   "DB611_Hydraulic_State_MH_Hydraulic{2}_Switch_Hydraulic_ON_OFF" : Bool = PLC DB939_Tool_alloc_HMI.SaveSortProg_name[7] AT %DB611.DBX26.3, 1 s
   "DB619_State_MPart_Recirculation{2}_Switch_Intervall" : Bool = PLC DB619_State_MPart.Recirculation[2].Switch_Intervall AT %DB619.DBX72.0, 1 s
   "DB619_State_MPart_Recirculation{2}_Switch_Lowpressure" : Bool = PLC DB619_State_MPart.Recirculation[2].Switch_Lowpressure AT %DB619.DBX72.2, 1 s
   "DB619_State_MPart_Recirculation{2}_Switch_Reduced" : Bool = PLC DB619_State_MPart.Recirculation[2].Switch_Reduced AT %DB619.DBX72.3, 1 s
   "DB619_State_MPart_Recirculation{2}_State_Intervall" : Int = PLC DB619_State_MPart.Recirculation[2].State_Intervall AT %DB619.DBW74, 1 s
   "DB619_State_MPart_Recirculation{2}_State_Lowpressure" : Int = PLC DB619_State_MPart.Recirculation[2].State_Lowpressure AT %DB619.DBW76, 1 s
   "DB619_State_MPart_Recirculation{2}_State_Reduced" : Int = PLC DB619_State_MPart.Recirculation[2].State_Reduced AT %DB619.DBW78, 1 s

HMI tags "General Machine Configuration"
   "DB790_PlantParameter_AmountMH" : Int = PLC DB790_PlantParameter.AmountMH AT %DB790.DBW4, 1 s
   "DB790_PlantParameter_AmountTank" : Int = PLC DB790_PlantParameter.AmountTank AT %DB790.DBW6, 1 s
   "DB790_PlantParameter_AmountToolStation" : Int = PLC DB790_PlantParameter.AmountToolStation AT %DB790.DBW10, 1 s
   "DB790_PlantParameter_AmountMouldCarrier" : Int = PLC DB790_PlantParameter.AmountMouldCarrier AT %DB790.DBW12, 1 s
   "DB790_PlantParameter_AmountProCanModul" : Int = PLC DB790_PlantParameter.AmountProCanModul AT %DB790.DBW2, 1 s
   "DB790_PlantParameter_AmountMeteringUnits" : Int = PLC DB790_PlantParameter.AmountMeteringUnits AT %DB790.DBW8, 1 s
   "DB790_PlantParameter_AmountMachine" : Int = PLC DB790_PlantParameter.AmountMachine AT %DB790.DBW24, 1 s
   "DB790_PlantParameter_Bit_ProgrammNofromInterface" : Bool = PLC DB790_PlantParameter.Bit.ProgrammNofromInterface AT %DB790.DBX0.3, 1 s
   "DB790_PlantParameter_Bit_MHNofromInterface" : Bool = PLC DB790_PlantParameter.Bit.MHNofromInterface AT %DB790.DBX0.2, 1 s
   "DB790_PlantParameter_AmountRobots" : Int = PLC DB790_PlantParameter.AmountRobots AT %DB790.DBW26, 1 s

HMI tags "Pump"
   "DB608_PV_Metering_Metering{0}_MixingRatio_PV_SetV_WarningLowerLimit" : Real = PLC DB608_PV_Metering.Metering[0].MixingRatio.PV_SetV.WarningLowerLimit AT %DB608.DBD202, 1 s
      on ChangeValue: SetBit("DB608_PV_Metering_Write")
   "DB608_PV_Metering_Metering{0}_MixingRatio_PV_SetV_WarningUpperLimit" : Real = PLC DB608_PV_Metering.Metering[0].MixingRatio.PV_SetV.WarningUpperLimit AT %DB608.DBD206, 1 s
      on ChangeValue: SetBit("DB608_PV_Metering_Write")
   "DB608_PV_Metering_Metering{0}_MixingRatio_PV_SetV_AlarmLowerLimit" : Real = PLC DB608_PV_Metering.Metering[0].MixingRatio.PV_SetV.AlarmLowerLimit AT %DB608.DBD210, 1 s
      on ChangeValue: SetBit("DB608_PV_Metering_Write")
   "DB608_PV_Metering_Metering{0}_MixingRatio_PV_SetV_AlarmUpperLimit" : Real = PLC DB608_PV_Metering.Metering[0].MixingRatio.PV_SetV.AlarmUpperLimit AT %DB608.DBD214, 1 s
      on ChangeValue: SetBit("DB608_PV_Metering_Write")
   "DB608_PV_Metering_Metering{0}_MixingRatio_PV_SetV_Value" : Real = PLC DB608_PV_Metering.Metering[0].MixingRatio.PV_SetV.Value AT %DB608.DBD198, 1 s
      on ChangeValue: SetBit("DB608_PV_Metering_Write")
   "DB608_PV_Metering_Metering{0}_Flow_PV_SetV_Value" : Real = PLC DB608_PV_Metering.Metering[0].Flow.PV_SetV.Value AT %DB608.DBD6, 1 s
      on ChangeValue: SetBit("DB608_PV_Metering_Write")
   "DB608_PV_Metering_Metering{0}_Flow_PV_SetV_WarningLowerLimit" : Real = PLC DB608_PV_Metering.Metering[0].Flow.PV_SetV.WarningLowerLimit AT %DB608.DBD10, 1 s
      on ChangeValue: SetBit("DB608_PV_Metering_Write")
   "DB608_PV_Metering_Metering{0}_Flow_PV_SetV_WarningUpperLimit" : Real = PLC DB608_PV_Metering.Metering[0].Flow.PV_SetV.WarningUpperLimit AT %DB608.DBD14, 1 s
      on ChangeValue: SetBit("DB608_PV_Metering_Write")
   "DB608_PV_Metering_Metering{0}_Flow_PV_SetV_AlarmLowerLimit" : Real = PLC DB608_PV_Metering.Metering[0].Flow.PV_SetV.AlarmLowerLimit AT %DB608.DBD18, 1 s
      on ChangeValue: SetBit("DB608_PV_Metering_Write")
   "DB608_PV_Metering_Metering{0}_Flow_PV_SetV_AlarmUpperLimit" : Real = PLC DB608_PV_Metering.Metering[0].Flow.PV_SetV.AlarmUpperLimit AT %DB608.DBD22, 1 s
      on ChangeValue: SetBit("DB608_PV_Metering_Write")
   "DB608_PV_Metering_Metering{0}_Pressure_PV_SetV_Value" : Real = PLC DB608_PV_Metering.Metering[0].Pressure.PV_SetV.Value AT %DB608.DBD54, 1 s
      on ChangeValue: SetBit("DB608_PV_Metering_Write")
   "DB608_PV_Metering_Metering{0}_Pressure_PV_SetV_WarningLowerLimit" : Real = PLC DB608_PV_Metering.Metering[0].Pressure.PV_SetV.WarningLowerLimit AT %DB608.DBD58, 1 s
      on ChangeValue: SetBit("DB608_PV_Metering_Write")
   "DB608_PV_Metering_Metering{0}_Pressure_PV_SetV_WarningUpperLimit" : Real = PLC DB608_PV_Metering.Metering[0].Pressure.PV_SetV.WarningUpperLimit AT %DB608.DBD62, 1 s
      on ChangeValue: SetBit("DB608_PV_Metering_Write")
   "DB608_PV_Metering_Metering{0}_Pressure_PV_SetV_AlarmLowerLimit" : Real = PLC DB608_PV_Metering.Metering[0].Pressure.PV_SetV.AlarmLowerLimit AT %DB608.DBD66, 1 s
      on ChangeValue: SetBit("DB608_PV_Metering_Write")
   "DB608_PV_Metering_Metering{0}_Pressure_PV_SetV_AlarmUpperLimit" : Real = PLC DB608_PV_Metering.Metering[0].Pressure.PV_SetV.AlarmUpperLimit AT %DB608.DBD70, 1 s
      on ChangeValue: SetBit("DB608_PV_Metering_Write")
   "Metering Display Open" : Int AT %DB1.DBD0
   "DB613_Komponent_State_Read" : Bool = PLC DB613_Komponent_State.Read AT %DB613.DBX6.0, 1 s
   "DB608_PV_Metering_Write" : Bool = PLC DB608_PV_Metering.Write AT %DB608.DBX4.1, 1 s
   "DB613_Komponent_State_ReadDeviceNo" : Int = PLC DB613_Komponent_State.ReadDeviceNo AT %DB613.DBW0, 1 s
      on ChangeValue: SetBit("DB613_Komponent_State_Write")
   "Control" : Int AT %DB1.DBW0
   "DB753_MeteringPump_Pump{0}_MachineNumber" : Byte = PLC DB753_MeteringPump.Pump[0].MachineNumber AT %DB753.DBB25, 1 s
      on ChangeValue: SetBit("DB613_Komponent_State_Write")
   "DB753_MeteringPump_Pump{0}_Name" : String[20] = PLC DB753_MeteringPump.Pump[0].Name AT %DB753.DBX26.0, 1 s
      on ChangeValue: SetBit("DB613_Komponent_State_Write")
   "DB753_MeteringPump_Pump{0}_TankNo" : Int = PLC DB753_MeteringPump.Pump[0].TankNo AT %DB753.DBW48, 1 s
      on ChangeValue: SetBit("DB613_Komponent_State_Write")
   "DB753_MeteringPump_Pump{0}_Pulse_per_liter" : Real = PLC DB753_MeteringPump.Pump[0].Pulse_per_liter AT %DB753.DBD52, 1 s
      on ChangeValue: SetBit("DB613_Komponent_State_Write")
   "DB753_MeteringPump_Pump{0}_MaxFlowLiter" : Real = PLC DB753_MeteringPump.Pump[0].MaxFlowLiter AT %DB753.DBD56, 1 s
      on ChangeValue: SetTag("DB613_Komponent_State_Write", 0)
   "DB753_MeteringPump_Pump{0}_MinFlowPercent" : Real = PLC DB753_MeteringPump.Pump[0].MinFlowPercent AT %DB753.DBD60, 1 s
      on ChangeValue: SetBit("DB613_Komponent_State_Write")
   "DB753_MeteringPump_Pump{0}_MaxFlowPercent" : Real = PLC DB753_MeteringPump.Pump[0].MaxFlowPercent AT %DB753.DBD64, 1 s
      on ChangeValue: SetBit("DB613_Komponent_State_Write")
   "DB753_MeteringPump_Pump{0}_Pump_Active" : Bool = PLC DB753_MeteringPump.Pump[0].Pump_Active AT %DB753.DBX22.0, 1 s
      on ChangeValue: SetBit("DB613_Komponent_State_Write")
   "DB753_MeteringPump_Pump{0}_WithFC" : Bool = PLC DB753_MeteringPump.Pump[0].WithFC AT %DB753.DBX22.1, 1 s
      on ChangeValue: SetBit("DB613_Komponent_State_Write")
   "DB753_MeteringPump_Pump{0}_With_2Point" : Bool = PLC DB753_MeteringPump.Pump[0].With_2Point AT %DB753.DBX22.2, 1 s
      on ChangeValue: SetBit("DB613_Komponent_State_Write")
   "DB753_MeteringPump_Pump{0}_WithFlowControl" : Bool = PLC DB753_MeteringPump.Pump[0].WithFlowControl AT %DB753.DBX22.3, 1 s
      on ChangeValue: SetBit("DB613_Komponent_State_Write")
   "DB753_MeteringPump_Pump{0}_WithoutFlowControl" : Bool = PLC DB753_MeteringPump.Pump[0].WithoutFlowControl AT %DB753.DBX22.4, 1 s
      on ChangeValue: SetBit("DB613_Komponent_State_Write")
   "DB753_MeteringPump_Pump{0}_WithFeedPump" : Bool = PLC DB753_MeteringPump.Pump[0].WithFeedPump AT %DB753.DBX22.5, 1 s
      on ChangeValue: SetBit("DB613_Komponent_State_Write")
   "DB753_MeteringPump_Pump{0}_WithEdgeFilter" : Bool = PLC DB753_MeteringPump.Pump[0].WithEdgeFilter AT %DB753.DBX22.6, 1 s
      on ChangeValue: SetBit("DB613_Komponent_State_Write")
   "DB753_MeteringPump_Pump{0}_PumDeselectionEnable" : Bool = PLC DB753_MeteringPump.Pump[0].PumDeselectionEnable AT %DB753.DBX22.7, 1 s
      on ChangeValue: SetBit("DB613_Komponent_State_Write")
   "DB753_MeteringPump_Pump{0}_PumpDeselected" : Bool = PLC DB753_MeteringPump.Pump[0].PumpDeselected AT %DB753.DBX23.0, 1 s
      on ChangeValue: SetBit("DB613_Komponent_State_Write")
   "DB753_MeteringPump_Pump{0}_PumpDeselectedInterval" : Bool = PLC DB753_MeteringPump.Pump[0].PumpDeselectedInterval AT %DB753.DBX23.1, 1 s
      on ChangeValue: SetBit("DB613_Komponent_State_Write")
   "DB753_MeteringPump_Pump{0}_WithFischerValveHP" : Bool = PLC DB753_MeteringPump.Pump[0].WithFischerValveHP AT %DB753.DBX23.2, 1 s
      on ChangeValue: SetBit("DB613_Komponent_State_Write")
   "DB753_MeteringPump_Pump{0}_WithFischerValveLP" : Bool = PLC DB753_MeteringPump.Pump[0].WithFischerValveLP AT %DB753.DBX23.3, 1 s
      on ChangeValue: SetBit("DB613_Komponent_State_Write")
   "DB753_MeteringPump_Pump{0}_WithHPHeatExchanger" : Bool = PLC DB918_ShotResultlast10.FilteredShot[6].Name[2] AT %DB753.DBX23.4, 1 s
      on ChangeValue: SetBit("DB613_Komponent_State_Write")
   "DB753_MeteringPump_Pump{0}_WithLPHeatExchanger" : Bool = PLC DB753_MeteringPump.Pump[0].WithLPHeatExchanger AT %DB753.DBX23.5, 1 s
      on ChangeValue: SetBit("DB613_Komponent_State_Write")
   "DB753_MeteringPump_Pump{0}_WithExhauseSystem" : Bool = PLC DB753_MeteringPump.Pump[0].WithExhauseSystem AT %DB753.DBX23.6, 1 s
      on ChangeValue: SetBit("DB613_Komponent_State_Write")
   "DB753_MeteringPump_Pump{0}_WithHeating" : Bool = PLC DB753_MeteringPump.Pump[0].WithHeating AT %DB753.DBX23.7, 1 s
      on ChangeValue: SetBit("DB613_Komponent_State_Write")
   "DB753_MeteringPump_Pump{0}_WithPipeHeating" : Bool = PLC DB918_ShotResultlast10.FilteredShot[6].MaterialConsumption[2] AT %DB753.DBX24.0, 1 s
      on ChangeValue: SetBit("DB613_Komponent_State_Write")
   "DB753_MeteringPump_Pump{0}_WithMinTempRelease" : Bool = PLC DB753_MeteringPump.Pump[0].WithMinTempRelease AT %DB753.DBX24.1, 1 s
      on ChangeValue: SetBit("DB613_Komponent_State_Write")
   "DB753_MeteringPump_Pump{0}_WithFlowFactor" : Bool = PLC DB753_MeteringPump.Pump[0].WithFlowFactor AT %DB753.DBX24.2, 1 s
      on ChangeValue: SetBit("DB613_Komponent_State_Write")
   "DB753_MeteringPump_Pump{0}_With_1Speed" : Bool = PLC DB753_MeteringPump.Pump[0].With_1Speed AT %DB753.DBX24.3, 1 s
      on ChangeValue: SetBit("DB613_Komponent_State_Write")
   "DB753_MeteringPump_Pump{0}_With_2Speed" : Bool = PLC DB753_MeteringPump.Pump[0].With_2Speed AT %DB753.DBX24.4, 1 s
      on ChangeValue: SetBit("DB613_Komponent_State_Write")
   "DB753_MeteringPump_Pump{0}_WithExternalFan" : Bool = PLC DB753_MeteringPump.Pump[0].WithExternalFan AT %DB753.DBX24.5, 1 s
      on ChangeValue: SetBit("DB613_Komponent_State_Write")
   "Control2" : Int, internal
   "OpenPidDialog" : Int, internal
   "DB613_Komponent_State_Write" : Bool = PLC DB613_Komponent_State.Write AT %DB613.DBX6.1, 1 s
   "DB751_auxiliaryDriveMetering_FeedingPumpControler{0}_ProportionalGain" : Real = PLC DB751_auxiliaryDriveMetering.FeedingPumpControler[0].ProportionalGain AT %DB701.DBD942, 1 s
      on ChangeValue: SetBit("DB613_Komponent_State_Write")
   "DB751_auxiliaryDriveMetering_FeedingPumpControler{0}_ResetTime" : Real = PLC DB751_auxiliaryDriveMetering.FeedingPumpControler[0].ResetTime AT %DB701.DBD946, 1 s
      on ChangeValue: SetBit("DB613_Komponent_State_Write")
   "DB751_auxiliaryDriveMetering_FeedingPumpControler{0}_DerivativeTime" : Real = PLC DB751_auxiliaryDriveMetering.FeedingPumpControler[0].DerivativeTime AT %DB701.DBD950, 1 s
      on ChangeValue: SetBit("DB613_Komponent_State_Write")
   "DB753_MeteringPump_Pump{0}_FlowFactor" : Real = PLC DB753_MeteringPump.Pump[0].FlowFactor AT %DB753.DBD72, 1 s
      on ChangeValue: SetBit("DB613_Komponent_State_Write")
   "DB753_MeteringPump_Pump{0}_DelayPressureFeedP" : S5Time = PLC DB753_MeteringPump.Pump[0].DelayPressureFeedP AT %DB753.DBW14, 1 s
      on ChangeValue: SetBit("DB613_Komponent_State_Write")
   "DB753_MeteringPump_Pump{0}_DelayRunTimeFeedP" : S5Time = PLC DB753_MeteringPump.Pump[0].DelayRunTimeFeedP AT %DB753.DBW16, 1 s
      on ChangeValue: SetBit("DB613_Komponent_State_Write")
   "DB751_auxiliaryDriveMetering_FeedingPump{0}_RunTime" : S5Time = PLC DB751_auxiliaryDriveMetering.FeedingPump[0].RunTime AT %DB701.DBW8, 1 s
      on ChangeValue: SetBit("DB613_Komponent_State_Write")
   "DB751_auxiliaryDriveMetering_FeedingPump{0}_PauseTime" : S5Time = PLC DB751_auxiliaryDriveMetering.FeedingPump[0].PauseTime AT %DB701.DBW10, 1 s
      on ChangeValue: SetBit("DB613_Komponent_State_Write")
   "DB751_auxiliaryDriveMetering_FeedingPump{0}_MinTempRelease" : Int = PLC DB751_auxiliaryDriveMetering.FeedingPump[0].MinTempRelease AT %DB701.DBW12, 1 s
      on ChangeValue: SetBit("DB613_Komponent_State_Write")
   "DB751_auxiliaryDriveMetering_FeedingPump{0}_Config_Exist" : Bool = PLC DB751_auxiliaryDriveMetering.FeedingPump[0].Config_Exist AT %DB701.DBX6.0, 1 s
      on ChangeValue: SetBit("DB613_Komponent_State_Write")
   "DB751_auxiliaryDriveMetering_EdgeFilter{0}_RunTime" : S5Time = PLC DB751_auxiliaryDriveMetering.EdgeFilter[0].RunTime AT %DB701.DBW112, 1 s
      on ChangeValue: SetBit("DB613_Komponent_State_Write")
   "DB751_auxiliaryDriveMetering_EdgeFilter{0}_PauseTime" : S5Time = PLC DB751_auxiliaryDriveMetering.EdgeFilter[0].PauseTime AT %DB701.DBW114, 1 s
      on ChangeValue: SetBit("DB613_Komponent_State_Write")
   "DB608_PV_Metering_HeatexchangerHP{0}_PV_SetV_Value" : Real = PLC DB608_PV_Metering.HeatexchangerHP[0].PV_SetV.Value AT %DB608.DBD3126, 1 s
      on ChangeValue: SetBit("DB613_Komponent_State_Write")
   "DB608_PV_Metering_HeatexchangerLP{0}_PV_SetV_Value" : Real = PLC DB608_PV_Metering.HeatexchangerLP[0].PV_SetV.Value AT %DB608.DBD3750, 1 s
      on ChangeValue: SetBit("DB613_Komponent_State_Write")
   "DB753_MeteringPump_Pump{0}_MinTempRelease" : Real = PLC DB753_MeteringPump.Pump[0].MinTempRelease AT %DB753.DBD18, 1 s
      on ChangeValue: SetBit("DB613_Komponent_State_Write")
   "DB613_Komponent_State_FeedPump{0}_Switch_Drive_ON_OFF" : Bool = PLC DB613_Komponent_State.FeedPump[0].Switch_Drive_ON_OFF AT %DB613.DBX61.3, 1 s
      on ChangeValue: SetBit("DB613_Komponent_State_Write")
   "DB613_Komponent_State_EdgeFilter{0}_Switch_Drive_ON_OFF" : Bool = PLC DB613_Komponent_State.EdgeFilter[0].Switch_Drive_ON_OFF AT %DB613.DBX9.7, 1 s
      on ChangeValue: SetBit("DB613_Komponent_State_Write")
   "DB613_Komponent_State_HeatexchangerHP{0}_Switch_Temp_ON_OFF" : Bool = PLC DB613_Komponent_State.HeatexchangerHP[0].Switch_Temp_ON_OFF AT %DB613.DBX763.7, 1 s
      on ChangeValue: SetBit("DB613_Komponent_State_Write")
   "DB613_Komponent_State_HeatexchangerLP{0}_Switch_Temp_ON_OFF" : Bool = PLC DB613_Komponent_State.HeatexchangerLP[0].Switch_Temp_ON_OFF AT %DB613.DBX867.7, 1 s
      on ChangeValue: SetBit("DB613_Komponent_State_Write")
   "DB613_Komponent_State_ActualDeviceNo" : Int = PLC DB613_Komponent_State.ActualDeviceNo AT %DB613.DBW2, 1 s
      on ChangeValue: SetBit("DB613_Komponent_State_Write")
   "DB753_MeteringPump_Pump{2}_Name" : String[20] = PLC DB753_MeteringPump.Pump[2].Name AT %DB753.DBX166.0, 1 s
   "DB753_MeteringPump_Pump{1}_Name" : String[20] = PLC DB753_MeteringPump.Pump[1].Name AT %DB753.DBX96.0, 1 s
   "DB608_PV_Metering_Read" : Bool = PLC DB608_PV_Metering.Read AT %DB608.DBX4.0, 1 s
   "DB753_MeteringPump_Pump{3}_Name" : String[20] = PLC DB753_MeteringPump.Pump[3].Name AT %DB753.DBX236.0, 1 s
   "DB753_MeteringPump_Pump{4}_Name" : String[20] = PLC DB753_MeteringPump.Pump[4].Name AT %DB753.DBX306.0, 1 s
   "DB753_MeteringPump_Pump{5}_Name" : String[20] = PLC DB753_MeteringPump.Pump[5].Name AT %DB753.DBX376.0, 1 s
   "DB753_MeteringPump_Pump{6}_Name" : String[20] = PLC DB753_MeteringPump.Pump[6].Name AT %DB753.DBX446.0, 1 s
   "DB753_MeteringPump_Pump{7}_Name" : String[20] = PLC DB753_MeteringPump.Pump[7].Name AT %DB753.DBX516.0, 1 s
   "DB753_MeteringPump_Pump{8}_Name" : String[20] = PLC DB753_MeteringPump.Pump[8].Name AT %DB753.DBX586.0, 1 s
   "DB753_MeteringPump_Pump{9}_Name" : String[20] = PLC DB753_MeteringPump.Pump[9].Name AT %DB753.DBX656.0, 1 s
   "DB753_MeteringPump_Pump{10}_Name" : String[20] = PLC DB753_MeteringPump.Pump[10].Name AT %DB753.DBX726.0, 1 s
   "DB753_MeteringPump_Pump{11}_Name" : String[20] = PLC DB753_MeteringPump.Pump[11].Name AT %DB753.DBX796.0, 1 s
   "DB753_MeteringPump_Pump{12}_Name" : String[20] = PLC DB753_MeteringPump.Pump[12].Name AT %DB753.DBX866.0, 1 s
   "DB613_Komponent_State_GroupStatus{1}_FaultExist" : Bool = PLC DB613_Komponent_State.GroupStatus[1].FaultExist AT %DB613.DBX739.0, 1 s
   "DB613_Komponent_State_GroupStatus{2}_FaultExist" : Bool = PLC DB613_Komponent_State.GroupStatus[2].FaultExist AT %DB613.DBX741.0, 1 s
   "DB751_auxiliaryDriveMetering_EdgeFilter{0}_Config_Driven" : Bool = PLC DB751_auxiliaryDriveMetering.EdgeFilter[0].Config_Driven AT %DB701.DBX110.1, 1 s
      on ChangeValue: SetBit("DB613_Komponent_State_Write")
   "DB751_auxiliaryDriveMetering_EdgeFilter{0}_Config_Double" : Bool = PLC DB751_auxiliaryDriveMetering.EdgeFilter[0].Config_Double AT %DB701.DBX110.3, 1 s
      on ChangeValue: SetBit("DB613_Komponent_State_Write")
   "DB751_auxiliaryDriveMetering_FeedingPump{0}_Config_With_PresControl" : Bool = PLC DB751_auxiliaryDriveMetering.FeedingPump[0].Config_With_PresControl AT %DB701.DBX6.3, 1 s
      on ChangeValue: SetBit("DB613_Komponent_State_Write")
   "DB751_auxiliaryDriveMetering_FeedingPump{0}_Config_WithFC" : Bool = PLC DB751_auxiliaryDriveMetering.FeedingPump[0].Config_WithFC AT %DB701.DBX6.1, 1 s
      on ChangeValue: SetBit("DB613_Komponent_State_Write")
   "DB751_auxiliaryDriveMetering_FeedingPump{0}_Config_Without_PresControl" : Bool = PLC DB751_auxiliaryDriveMetering.FeedingPump[0].Config_Without_PresControl AT %DB701.DBX6.2, 1 s
      on ChangeValue: SetBit("DB613_Komponent_State_Write")
   "DB751_auxiliaryDriveMetering_FeedingPump{0}_Config_Bypass" : Bool = PLC DB751_auxiliaryDriveMetering.FeedingPump[0].Config_Bypass AT %DB701.DBX6.4, 1 s
      on ChangeValue: SetBit("DB613_Komponent_State_Write")
   "DB751_auxiliaryDriveMetering_FeedingPump{0}_Config_Filling" : Bool = PLC DB751_auxiliaryDriveMetering.FeedingPump[0].Config_Filling AT %DB701.DBX6.5, 1 s
      on ChangeValue: SetBit("DB613_Komponent_State_Write")
   "DB751_auxiliaryDriveMetering_FeedingPump{0}_Config_ManualSwitchON" : Bool = PLC DB751_auxiliaryDriveMetering.FeedingPump[0].Config_ManualSwitchON AT %DB701.DBX6.6, 1 s
      on ChangeValue: SetBit("DB613_Komponent_State_Write")
   "DB613_Komponent_State_FlowPumpMin{0}" : Real = PLC DB613_Komponent_State.FlowPumpMin[0] AT %DB613.DBD268, 1 s
   "DB613_Komponent_State_FlowPumpMax{0}" : Real = PLC DB613_Komponent_State.FlowPumpMax[0] AT %DB613.DBD320, 1 s
   "DB613_Komponent_State_EdgeFilter{0}_State_Drive" : Int = PLC DB613_Komponent_State.EdgeFilter[0].State_Drive AT %DB613.DBW10, 1 s
   "DB613_Komponent_State_FeedPump{0}_State_Drive" : Int = PLC DB613_Komponent_State.FeedPump[0].State_Drive AT %DB613.DBW64, 1 s
   "DB613_Komponent_State_HeatexchangerHP{0}_State_Temp" : Int = PLC DB613_Komponent_State.HeatexchangerHP[0].State_Temp AT %DB613.DBW768, 1 s
   "DB613_Komponent_State_HeatexchangerLP{0}_State_Temp" : Int = PLC DB613_Komponent_State.HeatexchangerLP[0].State_Temp AT %DB613.DBW872, 1 s
   "DB613_Komponent_State_FeedPump{0}_FLT_Exist" : Bool = PLC DB613_Komponent_State.FeedPump[0].FLT_Exist AT %DB613.DBX60.0, 1 s
   "DB613_Komponent_State_HeatexchangerHP{0}_Fault_Exist" : Bool = PLC DB613_Komponent_State.HeatexchangerHP[0].Fault_Exist AT %DB613.DBX763.2, 1 s
   "DB613_Komponent_State_EdgeFilter{0}_FLT_Exist" : Bool = PLC DB613_Komponent_State.EdgeFilter[0].FLT_Exist AT %DB613.DBX8.0, 1 s
   "DB613_Komponent_State_MeteringPump{0}_FLT_Exist" : Bool = PLC DB613_Komponent_State.MeteringPump[0].FLT_Exist AT %DB613.DBX138.0, 1 s
   "DB613_Komponent_State_HeatexchangerLP{0}_Fault_Exist" : Bool = PLC DB613_Komponent_State.HeatexchangerLP[0].Fault_Exist AT %DB613.DBX867.2, 1 s
   "DB608_PV_Metering_Metering{0}_Pre_Pressure_PV_SetV_Value" : Real = PLC DB608_PV_Metering.Metering[0].Pre_Pressure.PV_SetV.Value AT %DB608.DBD150, 1 s
      on ChangeValue: SetBit("DB608_PV_Metering_Write")
   "DB753_MeteringPump_Pump{1}_WithEdgeFilter" : Bool = PLC DB753_MeteringPump.Pump[1].WithEdgeFilter AT %DB753.DBX92.6, 1 s
   "DB753_MeteringPump_Pump{2}_WithEdgeFilter" : Bool = PLC DB753_MeteringPump.Pump[2].WithEdgeFilter AT %DB753.DBX162.6, 1 s
   "DB753_MeteringPump_Pump{2}_WithLPHeatExchanger" : Bool = PLC DB753_MeteringPump.Pump[2].WithLPHeatExchanger AT %DB753.DBX163.5, 1 s
   "DB753_MeteringPump_Pump{1}_WithLPHeatExchanger" : Bool = PLC DB753_MeteringPump.Pump[1].WithLPHeatExchanger AT %DB753.DBX93.5, 1 s
   "DB613_Komponent_State_FeedPump{0}_ManipValuePercent" : Int = PLC DB613_Komponent_State.FeedPump[0].ManipValuePercent AT %DB613.DBW62, 1 s
   "DB753_MeteringPump_Pump{1}_WithHeating" : Bool = PLC DB753_MeteringPump.Pump[1].WithHeating AT %DB753.DBX93.7, 1 s
   "DB753_MeteringPump_Pump{2}_WithHeating" : Bool = PLC DB753_MeteringPump.Pump[2].WithHeating AT %DB753.DBX163.7, 1 s

HMI tags "Osciloscope"
   "DB025_Oszilloskop_SkalierungGraphLinks_Startwert" : Int = PLC DB025_Oszilloskop.SkalierungGraphLinks.Startwert AT %DB25.DBW220, 1 s
   "DB025_Oszilloskop_SkalierungGraphLinks_Ebdwert" : Int = PLC DB025_Oszilloskop.SkalierungGraphLinks.Ebdwert AT %DB25.DBW222, 1 s
   "DB025_Oszilloskop_SkalierungGraphRechts_Startwert" : Int = PLC DB025_Oszilloskop.SkalierungGraphRechts.Startwert AT %DB25.DBW224, 1 s
   "DB025_Oszilloskop_SkalierungGraphRechts_Ebdwert" : Int = PLC DB025_Oszilloskop.SkalierungGraphRechts.Ebdwert AT %DB25.DBW226, 1 s
   "DB025_Oszilloskop_Graph{1}_Auswahl" : Int = PLC DB025_Oszilloskop.Graph[1].Auswahl AT %DB25.DBW0, 1 s
   "DB025_Oszilloskop_Graph{1}_Nummer" : Int = PLC DB025_Oszilloskop.Graph[1].Nummer AT %DB25.DBW2, 1 s
   "DB025_Oszilloskop_Graph{1}_Komponente" : Int = PLC DB025_Oszilloskop.Graph[1].Komponente AT %DB25.DBW4, 1 s
   "DB025_Oszilloskop_Graph{1}_Sensor" : Int = PLC DB025_Oszilloskop.Graph[1].Sensor AT %DB25.DBW6, 1 s
   "DB025_Oszilloskop_Graph{1}_Skalierung" : Real = PLC DB025_Oszilloskop.Graph[1].Skalierung AT %DB25.DBD12, 1 s
   "DB025_Oszilloskop_Graph{2}_Auswahl" : Int = PLC DB025_Oszilloskop.Graph[2].Auswahl AT %DB25.DBW22, 1 s
   "DB025_Oszilloskop_Graph{2}_Nummer" : Int = PLC DB025_Oszilloskop.Graph[2].Nummer AT %DB25.DBW24, 1 s
   "DB025_Oszilloskop_Graph{2}_Komponente" : Int = PLC DB025_Oszilloskop.Graph[2].Komponente AT %DB25.DBW26, 1 s
   "DB025_Oszilloskop_Graph{2}_Sensor" : Int = PLC DB025_Oszilloskop.Graph[2].Sensor AT %DB25.DBW28, 1 s
   "DB025_Oszilloskop_Graph{2}_Skalierung" : Real = PLC DB025_Oszilloskop.Graph[2].Skalierung AT %DB25.DBD34, 1 s
   "DB025_Oszilloskop_Graph{3}_Auswahl" : Int = PLC DB025_Oszilloskop.Graph[3].Auswahl AT %DB25.DBW44, 1 s
   "DB025_Oszilloskop_Graph{3}_Nummer" : Int = PLC DB025_Oszilloskop.Graph[3].Nummer AT %DB25.DBW46, 1 s
   "DB025_Oszilloskop_Graph{3}_Komponente" : Int = PLC DB025_Oszilloskop.Graph[3].Komponente AT %DB25.DBW48, 1 s
   "DB025_Oszilloskop_Graph{3}_Sensor" : Int = PLC DB025_Oszilloskop.Graph[3].Sensor AT %DB25.DBW50, 1 s
   "DB025_Oszilloskop_Graph{3}_Skalierung" : Real = PLC DB025_Oszilloskop.Graph[3].Skalierung AT %DB25.DBD56, 1 s
   "DB025_Oszilloskop_Graph{4}_Auswahl" : Int = PLC DB025_Oszilloskop.Graph[4].Auswahl AT %DB25.DBW66, 1 s
   "DB025_Oszilloskop_Graph{4}_Nummer" : Int = PLC DB025_Oszilloskop.Graph[4].Nummer AT %DB25.DBW68, 1 s
   "DB025_Oszilloskop_Graph{4}_Komponente" : Int = PLC DB025_Oszilloskop.Graph[4].Komponente AT %DB25.DBW70, 1 s
   "DB025_Oszilloskop_Graph{4}_Sensor" : Int = PLC DB025_Oszilloskop.Graph[4].Sensor AT %DB25.DBW72, 1 s
   "DB025_Oszilloskop_Graph{4}_Skalierung" : Real = PLC DB025_Oszilloskop.Graph[4].Skalierung AT %DB25.DBD78, 1 s
   "DB025_Oszilloskop_Graph{5}_Auswahl" : Int = PLC DB025_Oszilloskop.Graph[5].Auswahl AT %DB25.DBW88, 1 s
   "DB025_Oszilloskop_Graph{5}_Nummer" : Int = PLC DB025_Oszilloskop.Graph[5].Nummer AT %DB25.DBW90, 1 s
   "DB025_Oszilloskop_Graph{5}_Komponente" : Int = PLC DB025_Oszilloskop.Graph[5].Komponente AT %DB25.DBW92, 1 s
   "DB025_Oszilloskop_Graph{5}_Sensor" : Int = PLC DB025_Oszilloskop.Graph[5].Sensor AT %DB25.DBW94, 1 s
   "DB025_Oszilloskop_Graph{5}_Skalierung" : Real = PLC DB025_Oszilloskop.Graph[5].Skalierung AT %DB25.DBD100, 1 s
   "DB025_Oszilloskop_Graph{6}_Auswahl" : Int = PLC DB025_Oszilloskop.Graph[6].Auswahl AT %DB25.DBW110, 1 s
   "DB025_Oszilloskop_Graph{6}_Nummer" : Int = PLC DB025_Oszilloskop.Graph[6].Nummer AT %DB25.DBW112, 1 s
   "DB025_Oszilloskop_Graph{6}_Komponente" : Int = PLC DB025_Oszilloskop.Graph[6].Komponente AT %DB25.DBW114, 1 s
   "DB025_Oszilloskop_Graph{6}_Sensor" : Int = PLC DB025_Oszilloskop.Graph[6].Sensor AT %DB25.DBW116, 1 s
   "DB025_Oszilloskop_Graph{6}_Skalierung" : Real = PLC DB025_Oszilloskop.Graph[6].Skalierung AT %DB25.DBD122, 1 s
   "DB025_Oszilloskop_Graph{7}_Auswahl" : Int = PLC DB025_Oszilloskop.Graph[7].Auswahl AT %DB25.DBW132, 1 s
   "DB025_Oszilloskop_Graph{7}_Nummer" : Int = PLC DB025_Oszilloskop.Graph[7].Nummer AT %DB25.DBW134, 1 s
   "DB025_Oszilloskop_Graph{7}_Komponente" : Int = PLC DB025_Oszilloskop.Graph[7].Komponente AT %DB25.DBW136, 1 s
   "DB025_Oszilloskop_Graph{7}_Sensor" : Int = PLC DB025_Oszilloskop.Graph[7].Sensor AT %DB25.DBW138, 1 s
   "DB025_Oszilloskop_Graph{7}_Skalierung" : Real = PLC DB025_Oszilloskop.Graph[7].Skalierung AT %DB25.DBD144, 1 s
   "DB025_Oszilloskop_Graph{8}_Auswahl" : Int = PLC DB025_Oszilloskop.Graph[8].Auswahl AT %DB25.DBW154, 1 s
   "DB025_Oszilloskop_Graph{8}_Nummer" : Int = PLC DB025_Oszilloskop.Graph[8].Nummer AT %DB25.DBW156, 1 s
   "DB025_Oszilloskop_Graph{8}_Komponente" : Int = PLC DB025_Oszilloskop.Graph[8].Komponente AT %DB25.DBW158, 1 s
   "DB025_Oszilloskop_Graph{8}_Sensor" : Int = PLC DB025_Oszilloskop.Graph[8].Sensor AT %DB25.DBW160, 1 s
   "DB025_Oszilloskop_Graph{8}_Skalierung" : Real = PLC DB025_Oszilloskop.Graph[8].Skalierung AT %DB25.DBD166, 1 s
   "DB025_Oszilloskop_Graph{1}_Wert" : Real = PLC DB025_Oszilloskop.Graph[1].Wert AT %DB25.DBD16, 1 s
   "DB025_Oszilloskop_Graph{2}_Wert" : Real = PLC DB025_Oszilloskop.Graph[2].Wert AT %DB25.DBD38, 1 s
   "DB025_Oszilloskop_Graph{3}_Wert" : Real = PLC DB025_Oszilloskop.Graph[3].Wert AT %DB25.DBD60, 1 s
   "DB025_Oszilloskop_Graph{4}_Wert" : Real = PLC DB025_Oszilloskop.Graph[4].Wert AT %DB25.DBD82, 1 s
   "DB025_Oszilloskop_Graph{5}_Wert" : Real = PLC DB025_Oszilloskop.Graph[5].Wert AT %DB25.DBD104, 1 s
   "DB025_Oszilloskop_Graph{6}_Wert" : Real = PLC DB025_Oszilloskop.Graph[6].Wert AT %DB25.DBD126, 1 s
   "DB025_Oszilloskop_Graph{7}_Wert" : Real = PLC DB025_Oszilloskop.Graph[7].Wert AT %DB25.DBD148, 1 s
   "DB025_Oszilloskop_Graph{8}_Wert" : Real = PLC DB025_Oszilloskop.Graph[8].Wert AT %DB25.DBD170, 1 s

HMI tags "ShotCounterMixingHead"
   "DB_Zaehler_Anzeige_MH_Counter_Reset{1}" : Real = PLC DB_Zaehler_Anzeige.MH_Counter_Reset[1] AT %DB211.DBD508, 1 s
   "DB_Zaehler_Anzeige_MH_Counter_Reset{2}" : Real = PLC DB_Zaehler_Anzeige.MH_Counter_Reset[2] AT %DB211.DBD512, 1 s
   "DB_Zaehler_Anzeige_MH_Counter_Reset{3}" : Real = PLC DB_Zaehler_Anzeige.MH_Counter_Reset[3] AT %DB211.DBD516, 1 s
   "DB_Zaehler_Anzeige_MH_Counter_Reset{4}" : Real = PLC DB_Zaehler_Anzeige.MH_Counter_Reset[4] AT %DB211.DBD520, 1 s
   "DB_Zaehler_Anzeige_MH_Counter_Reset{5}" : Real = PLC DB_Zaehler_Anzeige.MH_Counter_Reset[5] AT %DB211.DBD524, 1 s
   "DB_Zaehler_Anzeige_MH_Counter_Reset{6}" : Real = PLC DB_Zaehler_Anzeige.MH_Counter_Reset[6] AT %DB211.DBD528, 1 s
   "DB_Zaehler_Anzeige_MH_Counter_Reset{7}" : Real = PLC DB_Zaehler_Anzeige.MH_Counter_Reset[7] AT %DB211.DBD532, 1 s
   "DB_Zaehler_Anzeige_MH_Counter_Reset{8}" : Real = PLC DB_Zaehler_Anzeige.MH_Counter_Reset[8] AT %DB211.DBD536, 1 s
   "DB_Zaehler_Anzeige_MH_Counter_Reset{9}" : Real = PLC DB_Zaehler_Anzeige.MH_Counter_Reset[9] AT %DB211.DBD540, 1 s
   "DB_Zaehler_Anzeige_MH_Counter_Reset{10}" : Real = PLC DB_Zaehler_Anzeige.MH_Counter_Reset[10] AT %DB211.DBD544, 1 s
   "DB_Zaehler_Anzeige_MH_Counter_PreShift{1}" : Real = PLC DB_Zaehler_Anzeige.MH_Counter_PreShift[1] AT %DB211.DBD444, 1 s
   "DB_Zaehler_Anzeige_MH_Counter_PreShift{2}" : Real = PLC DB_Zaehler_Anzeige.MH_Counter_PreShift[2] AT %DB211.DBD448, 1 s
   "DB_Zaehler_Anzeige_MH_Counter_PreShift{3}" : Real = PLC DB_Zaehler_Anzeige.MH_Counter_PreShift[3] AT %DB211.DBD452, 1 s
   "DB_Zaehler_Anzeige_MH_Counter_PreShift{4}" : Real = PLC DB_Zaehler_Anzeige.MH_Counter_PreShift[4] AT %DB211.DBD456, 1 s
   "DB_Zaehler_Anzeige_MH_Counter_PreShift{5}" : Real = PLC DB_Zaehler_Anzeige.MH_Counter_PreShift[5] AT %DB211.DBD460, 1 s
   "DB_Zaehler_Anzeige_MH_Counter_PreShift{6}" : Real = PLC DB_Zaehler_Anzeige.MH_Counter_PreShift[6] AT %DB211.DBD464, 1 s
   "DB_Zaehler_Anzeige_MH_Counter_PreShift{7}" : Real = PLC DB_Zaehler_Anzeige.MH_Counter_PreShift[7] AT %DB211.DBD468, 1 s
   "DB_Zaehler_Anzeige_MH_Counter_PreShift{8}" : Real = PLC DB_Zaehler_Anzeige.MH_Counter_PreShift[8] AT %DB211.DBD472, 1 s
   "DB_Zaehler_Anzeige_MH_Counter_PreShift{9}" : Real = PLC DB_Zaehler_Anzeige.MH_Counter_PreShift[9] AT %DB211.DBD476, 1 s
   "DB_Zaehler_Anzeige_MH_Counter_PreShift{10}" : Real = PLC DB_Zaehler_Anzeige.MH_Counter_PreShift[10] AT %DB211.DBD480, 1 s
   "DB_Zaehler_Anzeige_MH_Counter_ActualShift{1}" : Real = PLC DB_Zaehler_Anzeige.MH_Counter_ActualShift[1] AT %DB211.DBD380, 1 s
   "DB_Zaehler_Anzeige_MH_Counter_ActualShift{2}" : Real = PLC DB_Zaehler_Anzeige.MH_Counter_ActualShift[2] AT %DB211.DBD384, 1 s
   "DB_Zaehler_Anzeige_MH_Counter_ActualShift{3}" : Real = PLC DB_Zaehler_Anzeige.MH_Counter_ActualShift[3] AT %DB211.DBD388, 1 s
   "DB_Zaehler_Anzeige_MH_Counter_ActualShift{4}" : Real = PLC DB_Zaehler_Anzeige.MH_Counter_ActualShift[4] AT %DB211.DBD392, 1 s
   "DB_Zaehler_Anzeige_MH_Counter_ActualShift{5}" : Real = PLC DB_Zaehler_Anzeige.MH_Counter_ActualShift[5] AT %DB211.DBD396, 1 s
   "DB_Zaehler_Anzeige_MH_Counter_ActualShift{6}" : Real = PLC DB_Zaehler_Anzeige.MH_Counter_ActualShift[6] AT %DB211.DBD400, 1 s
   "DB_Zaehler_Anzeige_MH_Counter_ActualShift{7}" : Real = PLC DB_Zaehler_Anzeige.MH_Counter_ActualShift[7] AT %DB211.DBD404, 1 s
   "DB_Zaehler_Anzeige_MH_Counter_ActualShift{8}" : Real = PLC DB_Zaehler_Anzeige.MH_Counter_ActualShift[8] AT %DB211.DBD408, 1 s
   "DB_Zaehler_Anzeige_MH_Counter_ActualShift{9}" : Real = PLC DB_Zaehler_Anzeige.MH_Counter_ActualShift[9] AT %DB211.DBD412, 1 s
   "DB_Zaehler_Anzeige_MH_Counter_ActualShift{10}" : Real = PLC DB_Zaehler_Anzeige.MH_Counter_ActualShift[10] AT %DB211.DBD416, 1 s
   "DB_Zaehler_Anzeige_MH_Counter_NonReset{1}" : Real = PLC DB_Zaehler_Anzeige.MH_Counter_NonReset[1] AT %DB211.DBD572, 1 s
   "DB_Zaehler_Anzeige_MH_Counter_NonReset{2}" : Real = PLC DB_Zaehler_Anzeige.MH_Counter_NonReset[2] AT %DB211.DBD576, 1 s
   "DB_Zaehler_Anzeige_MH_Counter_NonReset{3}" : Real = PLC DB_Zaehler_Anzeige.MH_Counter_NonReset[3] AT %DB211.DBD580, 1 s
   "DB_Zaehler_Anzeige_MH_Counter_NonReset{4}" : Real = PLC DB_Zaehler_Anzeige.MH_Counter_NonReset[4] AT %DB211.DBD584, 1 s
   "DB_Zaehler_Anzeige_MH_Counter_NonReset{5}" : Real = PLC DB_Zaehler_Anzeige.MH_Counter_NonReset[5] AT %DB211.DBD588, 1 s
   "DB_Zaehler_Anzeige_MH_Counter_NonReset{6}" : Real = PLC DB_Zaehler_Anzeige.MH_Counter_NonReset[6] AT %DB211.DBD592, 1 s
   "DB_Zaehler_Anzeige_MH_Counter_NonReset{7}" : Real = PLC DB_Zaehler_Anzeige.MH_Counter_NonReset[7] AT %DB211.DBD596, 1 s
   "DB_Zaehler_Anzeige_MH_Counter_NonReset{8}" : Real = PLC DB_Zaehler_Anzeige.MH_Counter_NonReset[8] AT %DB211.DBD600, 1 s
   "DB_Zaehler_Anzeige_MH_Counter_NonReset{9}" : Real = PLC DB_Zaehler_Anzeige.MH_Counter_NonReset[9] AT %DB211.DBD604, 1 s
   "DB_Zaehler_Anzeige_MH_Counter_NonReset{10}" : Real = PLC DB_Zaehler_Anzeige.MH_Counter_NonReset[10] AT %DB211.DBD608, 1 s
   "DB_Zaehler_Anzeige_Read" : Bool = PLC DB_Zaehler_Anzeige.Read AT %DB211.DBX4.0, 1 s